FUNCTION "Wips Have Matching Index" : Bool   // FC111, SCL
{ S7_Optimized_Access := 'TRUE' }
VERSION : 0.1
   VAR_INPUT
      selected_station_wips : Array[0.."wipCount"] of "Station: Wip: Wip Module";
      evaluation_station_wips : Array[0.."wipCount"] of "Station: Wip: Wip Module";
   END_VAR
   VAR_TEMP
      code_selected : DInt;
      code_evaluation : DInt;
      p_selected : Int;
      p_evaluation : Int;
      ret : Bool;
   END_VAR
   VAR CONSTANT
      null_value : Int := -1;
   END_VAR
BEGIN
   REGION "SCAN EACH WIP IN SELECTED STATION"
       FOR #p_selected := 0 TO "wipCount" DO

           REGION "IGNORE EMPTY WIPS"
               IF #selected_station_wips[#p_selected].wip.code <> #null_value THEN

                   REGION "SCAN EACH WIP IN EVALUATION STATION"
                       FOR #p_evaluation := 0 TO "wipCount" DO

                           REGION "SAVE CODES TO LOCAL VARIABLES"
                               #code_selected := #selected_station_wips[#p_selected].wip.code;
                               #code_evaluation := #evaluation_station_wips[#p_evaluation].wip.code;
                           END_REGION

                           REGION "COMPARE CODES"
                               IF #code_selected = #code_evaluation THEN
                                   #ret := true;
                                   EXIT;
                               END_IF;
                           END_REGION

                       END_FOR;
                   END_REGION

                   REGION "EXIT OUTER LOOP IF FOUND"
                       IF #ret THEN
                           EXIT;
                       END_IF;
                   END_REGION

               END_IF;
           END_REGION

       END_FOR;
   END_REGION


   REGION "RETURN"
       #"Wips Have Matching Index" := #ret;
   END_REGION
END_FUNCTION

FUNCTION "Modify Selectable Station List: Matching WIP" : Void   // FC112, SCL
{ S7_Optimized_Access := 'TRUE' }
VERSION : 0.1
   VAR_INPUT
      saved_wips : Array[0.."hmi_station_count"] of "WIP: Station";
      selection_change : "Station Selection Change";
      selected_stations : "Selected Stations";
   END_VAR
   VAR_IN_OUT
      selectable_stns : Array[0.."stnCount"] of Int;
      selectable_stn_cnt : Int;
      visible_stations : Array[0.."slct_stn_btn_count"] of Int;
   END_VAR
   VAR_TEMP
      has_matching_wip : Bool;
      i : Int;
      p_evaluation : Int;
      selected_station : "WIP: Station";
      selected_stations_count : Int;
      selected_stations_indices : Array[0.."stnCount"] of Int;
      station_index : Int;
      t_selectable_stns : Array[0.."stnCount"] of Int;
      t_selectable_stn_count : Int;
   END_VAR
   VAR CONSTANT
      null_value : Int := -1;
   END_VAR
BEGIN
   REGION "SET UP LOCALS"
       #t_selectable_stns := #selectable_stns;
       #t_selectable_stn_count := #selectable_stn_cnt;
       #selected_stations_count := "Count Selected Stations"(#selected_stations.stns);
       "List of Array of Bool Indices"(array_of_bool := #selected_stations.stns,
                                       list_of_indices => #selected_stations_indices);
   END_REGION


   REGION "CHECK EACH SELECTED STATION VS SELECTABLE STATIONS"
       FOR #i := 0 TO #selected_stations_count DO

           REGION "EXIT LOOP ON FIRST NULL"
               IF #selected_stations_indices[#i] = #null_value THEN
                   EXIT;
               END_IF;
           END_REGION

           REGION "GET SELECTED STATION DATA"
               #station_index := #selected_stations_indices[#i];
               #selected_station := "Get WIP Station by Global Index"(index := #station_index,
                                                                         recipe_stations := #saved_wips);
           END_REGION

           REGION "REMOVE STATIONS WITH NON-MATCHING WIP"
               FOR #p_evaluation := 0 TO "hmi_station_count" DO

                   REGION "DONT RUN IF SELECTED AND EVALUATION STATIONS MATCH"
                       IF #selected_station.pStn <> #saved_wips[#p_evaluation].pStn THEN

                           REGION "RUN IF EVALUATION STATION IS SELECTABLE"
                               IF "Is In Int Array"(array_of_int := #selectable_stns, search_term := #saved_wips[#p_evaluation].pStn) THEN

                                   REGION "REMOVE EVALUATION STATION FROM SELECTABLE LIST IF NO MATCHING WIPS"
                                       #has_matching_wip := "Wips Have Matching Index"(selected_station_wips := #selected_station.wip,
                                                                                       evaluation_station_wips := #saved_wips[#p_evaluation].wip);
                                       IF NOT #has_matching_wip THEN
                                           #t_selectable_stns[#p_evaluation] := #null_value;
                                       END_IF;
                                   END_REGION

                               END_IF;
                           END_REGION

                       END_IF;
                   END_REGION

               END_FOR;
           END_REGION

           REGION "COLLAPSE"
               "Collapse Int Array"(null_value := #null_value,
                                    int_array := #t_selectable_stns);
           END_REGION

       END_FOR;
   END_REGION


   REGION "GET COUNT"
       #t_selectable_stn_count := "Count Collapsed Int Array"(null_value := #null_value,
                                                              array := #t_selectable_stns);
   END_REGION


   REGION "RETURN"
       #selectable_stns := #t_selectable_stns;
       #selectable_stn_cnt := #t_selectable_stn_count;
       "Remap Int Array"(source_int_array := #t_selectable_stns,
                         destination_int_array := #visible_stations);

   END_REGION
END_FUNCTION

FUNCTION "Pop Up: Select Stations: Animations" : Void   // FC119, SCL
{ S7_Optimized_Access := 'TRUE' }
VERSION : 0.1
   VAR_INPUT
      all_stations : "Station: All Stations";
      selectable_stn_cnt : Int;
      selected_stns : "Selected Stations";
      visable_stns : Array[0.."slct_stn_btn_count"] of Int;
   END_VAR
   VAR_IN_OUT
      interface : "Select Station";
   END_VAR
   VAR_TEMP
      i : Int;
      t_interface : "Select Station";
   END_VAR
BEGIN
   REGION "COPY TO LOCAL"
       #t_interface := #interface;
   END_REGION


   REGION "ANIMATE CLOSE SCREEN BUTTON"
       #t_interface.close_screen.animate := "Animate Bool"(colorTrue := "BgLGr",
                                                           colorFalse := "BgLRd",
                                                           evalSignal := #t_interface.close_screen.actuate);
   END_REGION


   REGION "ANIMATE STATION SELECT BUTTONS"

       REGION "ACTUATE"
           FOR #i := 0 TO "slct_stn_btn_count" DO
               IF #visable_stns[#i] <> -1 THEN

                   REGION "NOT SELECTED"
                       IF NOT #selected_stns.stns[#visable_stns[#i]] THEN
                           #t_interface.stn_select_btns[#i].animate := "Animate Bool"(colorTrue := "BgLGr",
                                                                                      colorFalse := "BgGray",
                                                                                      evalSignal := #t_interface.stn_select_btns[#i].actuate);
                       END_IF;
                   END_REGION

                   REGION "SELECTED"
                       IF #selected_stns.stns[#visable_stns[#i]] THEN
                           #t_interface.stn_select_btns[#i].animate := "Animate Bool"(colorTrue := "BgLGr",
                                                                                      colorFalse := "BgLBl",
                                                                                      evalSignal := #t_interface.stn_select_btns[#i].actuate);
                       END_IF;
                   END_REGION

               END_IF;
           END_FOR;
       END_REGION

       REGION "ENABLE"
           FOR #i := 0 TO "slct_stn_btn_count" DO
               #t_interface.stn_select_btns[#i].enable := "Select Station Button Activation"(btn_index := #i,
                                                                                             selectable_stn_cnt := #selectable_stn_cnt);
           END_FOR;
       END_REGION

       REGION "VISIBLE"
           FOR #i := 0 TO "slct_stn_btn_count" DO
               #t_interface.stn_select_btns[#i].visible := "Select Station Button Activation"(btn_index := #i,
                                                                                              selectable_stn_cnt := #selectable_stn_cnt);
           END_FOR;
       END_REGION

       REGION "DISABLED"
           FOR #i := 0 TO "slct_stn_btn_count" DO
               #t_interface.stn_select_btns[#i].enable := TRUE;
           END_FOR;
           FOR #i := #selectable_stn_cnt TO "slct_stn_btn_count" DO
               #t_interface.stn_select_btns[#i].enable := FALSE;
           END_FOR;
       END_REGION

       REGION "POPULATE STATION NAMES"
           FOR #i := 0 TO "slct_stn_btn_count" DO
               IF #visable_stns[#i] <> -1 THEN
                   #t_interface.stn_select_btns[#i].label := "Populate Station Name"(lines := 2,
                                                                                     stn := #all_stations.stn[#visable_stns[#i]]);
               END_IF;
           END_FOR;
       END_REGION

   END_REGION


   REGION "ANIMATE NAV BAR"

       REGION "NOTES"
           // mapping is necessary because hmi faceplate data structures
           // cannot consist of embedded udts
       END_REGION

       REGION "MAP HMI TO PLC"
           "Nav Bar Data Map: HMI to PLC"(hmi := #t_interface.nav_bar_HMI,
                                          plc := #t_interface.nav_Bar_PLC);
       END_REGION

       REGION "ANIMATION CALLS"
           "Select Station Nav Bar Button Animation"(selectable_stations := #selectable_stn_cnt,
                                                     visible_rows := "slct_stn_btn_count",
                                                     button := #t_interface.nav_Bar_PLC.top);
           "Select Station Nav Bar Button Animation"(selectable_stations := #selectable_stn_cnt,
                                                     visible_rows := "slct_stn_btn_count",
                                                     button := #t_interface.nav_Bar_PLC.pageUp);
           "Select Station Nav Bar Button Animation"(selectable_stations := #selectable_stn_cnt,
                                                     visible_rows := "slct_stn_btn_count",
                                                     button := #t_interface.nav_Bar_PLC.lineUp);
           "Select Station Nav Bar Button Animation"(selectable_stations := #selectable_stn_cnt,
                                                     visible_rows := "slct_stn_btn_count",
                                                     button := #t_interface.nav_Bar_PLC.lineDown);
           "Select Station Nav Bar Button Animation"(selectable_stations := #selectable_stn_cnt,
                                                     visible_rows := "slct_stn_btn_count",
                                                     button := #t_interface.nav_Bar_PLC.pageDown);
           "Select Station Nav Bar Button Animation"(selectable_stations := #selectable_stn_cnt,
                                                     visible_rows := "slct_stn_btn_count",
                                                     button := #t_interface.nav_Bar_PLC.bottom);
       END_REGION

       REGION "MAP PLC TO HMI"
           "Nav Bar Data Map: PLC to HMI"(plc := #t_interface.nav_Bar_PLC,
                                          hmi := #t_interface.nav_bar_HMI);
       END_REGION

   END_REGION


   REGION "DRAW"
       #interface := #t_interface;
   END_REGION
END_FUNCTION

// folder: HMI: Warehouse/Pop Ups/Select WIP

FUNCTION_BLOCK "Pop Up: Select WIPs"   // FB28, SCL
{ S7_Optimized_Access := 'TRUE' }
VERSION : 0.1
   VAR_INPUT
      stations : "Station: All Stations";
      wip_stations : Array[0.."hmi_station_count"] of "WIP: Station";
   END_VAR
   VAR_IN_OUT
      interface : "Select WIP";
      meta_data : "Setting Meta Data";
   END_VAR
   VAR
      selectable_wips_count : Int;
   END_VAR
   VAR_TEMP
      t_interface : "Select WIP";
   END_VAR
   VAR CONSTANT
      null_value : Int := -1;
   END_VAR
BEGIN
   IF #meta_data.selection_change.selection_change THEN
       IF "Is HMI Station"(#stations.stn[#meta_data.selection_change.station_index]) THEN
           "Pop Up: Select WIPs: Build Selectable List"(meta_data := #meta_data,
                                                        selected_stations := #meta_data.selected_stns,
                                                        wip_stations := #wip_stations,
                                                        stations := #stations,
                                                        selectable_wips_count := #selectable_wips_count);
       END_IF;
   END_IF;
END_FUNCTION_BLOCK

FUNCTION "Pop Up: Select WIPs: Get Matching WIPs" : Void   // FC125, SCL
{ S7_Optimized_Access := 'TRUE' }
VERSION : 0.1
   VAR_INPUT
      outer_wips : Array[0.."wipCount"] of "Station: Wip: Wip Module";
      inner_wips : Array[0.."wipCount"] of "Station: Wip: Wip Module";
   END_VAR
   VAR_IN_OUT
      selectable_wips : "Selectable Wips";
      selectable_wips_count : Int;
   END_VAR
   VAR_TEMP
      i : Int;
      j : Int;
      t_selectable_wips : "Selectable Wips";
      t_selectable_wips_count : Int;
   END_VAR
BEGIN
   REGION "COPY TO LOCAL"
       #t_selectable_wips := #selectable_wips;
       #t_selectable_wips_count := 0;
   END_REGION

   REGION "COMPARE EACH WIP CODE IN OUTER LIST ..." 
       FOR #i := 0 TO "wipCount" DO

           REGION "LEAVE LOOP ON FIRST NULL"
               IF #outer_wips[#i].wip.code = "null_value" THEN
                   EXIT;
               END_IF;
           END_REGION

           REGION "WITH EACH IN INNER LIST AND ..."
               FOR #j := 0 TO "wipCount" DO

                   REGION "COPY MATCHES"
                       IF #outer_wips[#i].wip.code = #inner_wips[#j].wip.code THEN
                           #t_selectable_wips.wips[#t_selectable_wips_count] := #outer_wips[#i].wip.code;
                           #t_selectable_wips_count += 1;
                       END_IF;
                   END_REGION

               END_FOR;
           END_REGION

       END_FOR;
   END_REGION


   REGION "RETURN"
       #selectable_wips := #t_selectable_wips;
       #selectable_wips_count := #t_selectable_wips_count;
   END_REGION
END_FUNCTION

FUNCTION "Pop Up: Select WIPs: Build Selectable List" : Void   // FC128, SCL
{ S7_Optimized_Access := 'TRUE' }
VERSION : 0.1
   VAR_INPUT
      selected_stations : "Selected Stations";
      stations : "Station: All Stations";
      wip_stations : Array[0.."hmi_station_count"] of "WIP: Station";
   END_VAR
   VAR_IN_OUT
      meta_data : "Setting Meta Data";
      selectable_wips_count : Int;
   END_VAR
   VAR_TEMP
      global_index : Int;
      inner_wip_index : Int;
      outer_wip_index : Int;
      p_outer : Int;
      p_inner : Int;
      selected_station_count : Int;
      station : "WIP: Station";
      t_selectable_wips_count : Int;
   END_VAR
BEGIN
   REGION "INITIALIZE SELECTABLE WIPS"
       "Fill DInt Array"(int_in := -1,
                         array_out => #meta_data.selectable_wips.wips);
       #t_selectable_wips_count := 0;
   END_REGION


   REGION "Count Selected Stations"
       #selected_station_count := "Count Selected Stations"(#selected_stations.stns);
   END_REGION


   REGION "SINGLE STATION SELECTION"
       IF #selected_station_count = 1 THEN
           #global_index := "Get First Selected Station"(#selected_stations.stns);
           #outer_wip_index := "Get WIP Station Index by Global Index"(wip_stations := #wip_stations,
                                                                       global_index := #global_index);
           "Pop Up: Select WIPs: Map WIP Codes"(wip_station := #wip_stations[#outer_wip_index],
                                                selectable_wips := #meta_data.selectable_wips,
                                                selectable_wip_count := #t_selectable_wips_count);
       END_IF;
   END_REGION


   REGION "MULTI STATION SELECTION"
       IF #selected_station_count > 1 THEN
           REGION "FOR EACH STATION..."
               FOR #p_outer := 0 TO "stnCount" DO

                   REGION "IF THE STATION HAS BEEN SELECTED..."
                       IF #selected_stations.stns[#p_outer] THEN

                           REGION "GET THE WIP STATION INDEX"
                               #outer_wip_index := "Get WIP Station Index by Global Index"(wip_stations := #wip_stations,
                                                                                           global_index := #p_outer);
                           END_REGION

                           REGION "FOR EACH STATION AFTER THIS STATION..."
                               FOR #p_inner := #p_outer + 1 TO "stnCount" DO

                                   REGION "IF THE STATION HAS BEEN SELECTED"
                                       IF #selected_stations.stns[#p_inner] THEN

                                           REGION "GET THE WIP STATION INDEX"
                                               #inner_wip_index := "Get WIP Station Index by Global Index"(wip_stations := #wip_stations,
                                                                                                           global_index := #p_inner);
                                           END_REGION

                                           REGION "INSERT INTO SELECTABLE WIP ARRAY"
                                               "Pop Up: Select WIPs: Get Matching WIPs"(outer_wips := #wip_stations[#outer_wip_index].wip,
                                                                                        inner_wips := #wip_stations[#inner_wip_index].wip,
                                                                                        selectable_wips := #meta_data.selectable_wips,
                                                                                        selectable_wips_count := #t_selectable_wips_count);
                                           END_REGION

                                       END_IF;
                                   END_REGION

                               END_FOR;
                           END_REGION

                       END_IF;
                   END_REGION

               END_FOR;
           END_REGION
       END_IF;
   END_REGION


   REGION "RETURN"
       #selectable_wips_count := #t_selectable_wips_count;
   END_REGION
END_FUNCTION

FUNCTION "Pop Up: Select WIPs: Map WIP Codes" : Void   // FC129, SCL
{ S7_Optimized_Access := 'TRUE' }
VERSION : 0.1
   VAR_INPUT
      wip_station : "WIP: Station";
   END_VAR
   VAR_IN_OUT
      selectable_wips : "Selectable Wips";
      selectable_wip_count : Int;
   END_VAR
   VAR_TEMP
      i : Int;
      t_selectable_wips : "Selectable Wips";
      t_selectable_wip_count : Int;
   END_VAR
BEGIN
   REGION "COPY TO LOCAL"
       #t_selectable_wips := #selectable_wips;
       #t_selectable_wip_count := #selectable_wip_count;
   END_REGION


   REGION "MAP VALUES"
       FOR #i := 0 TO "wipCount" DO
           IF #wip_station.wip[#i].wip.code = "null_value" THEN
               EXIT;
           END_IF;
           #t_selectable_wips.wips[#i] := #wip_station.wip[#i].wip.code;
       END_FOR;
   END_REGION


   REGION "COUNT SELECTABLE WIPS"
       #t_selectable_wip_count := "Count Collapsed DInt Array"(null_value := INT_TO_DINT("null_value"),
                                                               array := #t_selectable_wips.wips);
   END_REGION


   REGION "RETURN"
       #selectable_wips := #t_selectable_wips;
       #selectable_wip_count := #t_selectable_wip_count;
   END_REGION
END_FUNCTION

// folder: HMI: Warehouse/RSP Simulation

FUNCTION_BLOCK "Sim: from Global"   // FB26, SCL
{ S7_Optimized_Access := 'TRUE' }
VERSION : 0.1
   VAR_INPUT
      stns : "Station: All Stations";
   END_VAR
   VAR_IN_OUT
      simStations : "Simulated Stations";
   END_VAR
   VAR
      old : Struct
         nextGrp : Bool;
         prevGrp : Bool;
      END_STRUCT;
   END_VAR
   VAR_TEMP
      animate : USInt;
      btnCount : Int;
      currentBtn : Bool;
      dzLabel : WString;
      firstStn : Int;
      i : Int;
      intBox : Int;
      j : Int;
      kp8Color : DWord;
      label : WString;
      oldBtn : Bool;
      pSim : Int;
      pStn : Int;
   END_VAR
   VAR CONSTANT
      space : WString := WSTRING#' ';
      lead0 : WString := WSTRING#'0';
      volvo16 : WString := WSTRING#'VOLVO 16';
   END_VAR
BEGIN
   REGION "COPY TO LOCAL"
       #firstStn := #simStations.firstStn;
   END_REGION

   REGION "RESOLVE STATION POINTER"

       REGION "PROCESS NEXT GROUP PRESS"

           REGION "COPY TO LOCAL"
               #currentBtn := #simStations.down.actuate;
               #oldBtn := #old.nextGrp;
           END_REGION

           REGION "FALLING EDGE OF NEXT GROUP"
               IF NOT #currentBtn AND #oldBtn THEN

                   REGION "INCREMENT FIRST STATION"
                       #firstStn += "simKP8Count";
                   END_REGION

                   REGION "UPPER LIMIT ROLL OVER"
                       IF #firstStn > "stnCount" THEN
                           #firstStn -= "stnCount" + 1;
                       END_IF;
                   END_REGION

               END_IF;
           END_REGION

           REGION "NEXT GROUP CHANGE DETECTION"
               #old.nextGrp := #currentBtn;
           END_REGION

       END_REGION

       REGION "PROCESS PREVIOUS GROUP PRESS"

           REGION "COPY TO LOCAL"
               #currentBtn := #simStations.up.actuate;
               #oldBtn := #old.prevGrp;
           END_REGION

           REGION "FALLING EDGE OF PREVIOUS GROUP"
               IF NOT #currentBtn AND #oldBtn THEN

                   REGION "DECREMENT FIRST STATION"
                       #firstStn -= "simKP8Count";
                   END_REGION

                   REGION "LOWER LIMIT ROLL OVER"
                       IF #firstStn < 0 THEN
                           #firstStn += "stnCount" + 1;
                       END_IF;
                   END_REGION

               END_IF;
           END_REGION

           REGION "PREVIOUS GROUP CHANGE DETECTION"
               #old.prevGrp := #currentBtn;
           END_REGION

       END_REGION

   END_REGION

   REGION "FOR EACH BUTTON"
       FOR #i := 0 TO 11 DO

           REGION "CALCULATE POINTER"
               #pStn := #i + #firstStn;
               #pSim := #i;
           END_REGION

           REGION "UPPER LIMIT ROLL OVER"
               IF #pStn > "stnCount" THEN
                   #pStn := #firstStn + #i - "stnCount" - 1;
               END_IF;
           END_REGION

           REGION "COPY TO LOCAL"
               #kp8Color := #stns.stn[#pStn].wipCmpts.ioData.kp8.tempOut;
           END_REGION

           REGION "LABEL STATIONS"

               REGION "DETERMINE LINE LABEL"
                   #label := #stns.stn[#pStn].id.lineName;
                   IF #label = #volvo16 THEN
                       #label := WSTRING#'V16';
                   END_IF;
               END_REGION

               REGION "DETERMINE DROP ZONE LABEL"
                   #intBox := USINT_TO_INT(#stns.stn[#pStn].id.dropZone);
                   IF #intBox <= 9 THEN
                       #dzLabel := CONCAT_WSTRING(IN1 := #lead0,
                                                  IN2 := "Strip Sign"(INT_TO_WSTRING(#intBox)));
                   END_IF;
                   IF #intBox >= 10 THEN
                       #dzLabel := "Strip Sign"(INT_TO_WSTRING(#intBox));
                   END_IF;
               END_REGION

               REGION "WRITE LABEL"
                   #label := CONCAT_WSTRING(IN1 := #label,
                                            IN2 := #space,
                                            IN3 := #dzLabel);
                   #simStations.me[#pSim].stn.label := #label;
               END_REGION

           END_REGION

           REGION "ANIMATE STATION LABEL"
               #simStations.me[#pSim].stn.animate := "BgGray";
           END_REGION

           REGION "FOR EACH BUTTON"
               FOR #j := 0 TO "btnCount" DO

                   REGION "COLOR BUTTONS"
                       #animate := "KP8 Driver: HMI Emulator: Animation"(kp8Color := #kp8Color,
                                                                btnNumber := #j);
                       #simStations.me[#pSim].btn.animate[#j] := #animate;
                   END_REGION

                   REGION "WRITE BUTTON LABELS"
                       #intBox := "Pointer Calc: KP8 Labels"(#j);
                       #label := "Strip Sign"(INT_TO_WSTRING(#intBox));
                       #simStations.me[#pSim].btn.labels[#j] := #label;
                   END_REGION

               END_FOR;
           END_REGION

       END_FOR;
   END_REGION

   REGION "SAVE FIRST STATION"
       #simStations.firstStn := #firstStn;
   END_REGION

   REGION "ANIMATE NEXT GROUP PRESS"
       #simStations.down.animate := "Animate Bool"(colorTrue := "BgLGr",
                                                   colorFalse := "BgGray",
                                                   evalSignal := #simStations.down.actuate);
   END_REGION

   REGION "ANIMATE PREV GROUP PARESS"
       #simStations.up.animate := "Animate Bool"(colorTrue := "BgLGr",
                                                 colorFalse := "BgGray",
                                                 evalSignal := #simStations.up.actuate);
   END_REGION
END_FUNCTION_BLOCK

FUNCTION "Sim: to Global" : Void   // FC23, SCL
{ S7_Optimized_Access := 'TRUE' }
VERSION : 0.1
   VAR_INPUT
      simStns : "Simulated Stations";
   END_VAR
   VAR_IN_OUT
      stations : "Station: All Stations";
   END_VAR
   VAR_TEMP
      i : Int;
      j : Int;
      pSim : Int;
      pStn : Int;
   END_VAR
BEGIN
   REGION "COPY TO LOCAL"
       // #btnCount := "btnCount";
       // #firstStn := #simStns.firstStn;
       // #simKP8Count := "simKP8Count";
       // #stnCount := "stnCount";
   END_REGION

   REGION "FOR EACH STATION"
       FOR #i := 0 TO "simKP8Count" DO

           REGION "CALCULATE POINTER"
               #pStn := #i + #simStns.firstStn;
               #pSim := #i;
           END_REGION

           REGION "UPPER LIMIT ROLL OVER"
               IF #pStn > "stnCount" THEN
                   #pStn := #simStns.firstStn + #i - "stnCount" - 1;
               END_IF;
           END_REGION

           REGION "COPY SIMULATED PRESSES"
               #stations.stn[#pStn].wipCmpts.ioData.kp8.input.%B1 := #simStns.me[#pSim].btn.actuate;
           END_REGION

       END_FOR;
   END_REGION
END_FUNCTION

FUNCTION "Sim: KP8 Animations" : Word   // FC84, SCL
{ S7_Optimized_Access := 'TRUE' }
VERSION : 0.1
   VAR_INPUT
      pbs : DWord;
   END_VAR
   VAR_TEMP
      ret : Word;
   END_VAR
BEGIN
   #"Sim: KP8 Animations".%B1 := #pbs.%B0;
   #"Sim: KP8 Animations".%B0 := #pbs.%B1;
END_FUNCTION

// folder: OBs

ORGANIZATION_BLOCK "Rack or station failure"   // OB86, LAD, RackStationFailure
{ S7_Optimized_Access := 'TRUE' }
VERSION : 0.1
   VAR_INPUT
      LADDR : Hw_Device;   // Hardware identifier
      Event_Class : Byte;   // Event class
      Fault_ID : Byte;   // Fault identifier
   END_VAR
BEGIN
END_ORGANIZATION_BLOCK

ORGANIZATION_BLOCK "Startup"   // OB100, LAD, Startup
TITLE = "Complete Restart"
{ S7_Optimized_Access := 'TRUE' }
VERSION : 0.1
   VAR_INPUT
      LostRetentive : Bool;   // True if retentive data are lost
      LostRTC : Bool;   // True if date and time are lost
   END_VAR
BEGIN

REGION Network 1 (SCL): HMI STATION INITIALIZATION
   "HMI Station Initialization"();
END_REGION
END_ORGANIZATION_BLOCK

ORGANIZATION_BLOCK "Programming error"   // OB121, LAD, ProgrammingError
{ S7_Optimized_Access := 'TRUE' }
VERSION : 0.1
   VAR_INPUT
      BlockNr : UInt;   // Number of causing block
      Reaction : USInt;   // 0:ignore, 1:substitute, 2:skip
      Fault_ID : Byte;   // Fault identifier
      BlockType : USInt;   // 16#01:OB, 16#02:FC, 16#03:FB, 16#04:SFC, 16#05:SFB, 16#06:DB: Type of block causing the error
      Area : USInt;   // Area where the error occured
      DBNr : DB_ANY;   // DB number if Area = DB or DI
      Csg_OBNr : OB_Any;   // Number of OB causing the error
      Csg_Prio : USInt;   // Priority of OB causing the error
      Width : USInt;   // 0:bit, 1:byte, 2:word, 3:dword, 4:lword
   END_VAR
BEGIN
END_ORGANIZATION_BLOCK

ORGANIZATION_BLOCK "IO access error"   // OB122, LAD, IOAccessError
{ S7_Optimized_Access := 'TRUE' }
VERSION : 0.1
   VAR_INPUT
      BlockNr : UInt;   // Number of causing block
      Reaction : USInt;   // 0:ignore, 1:substitute, 2:skip
      Fault_ID : Byte;   // 16#42:reading, 16#43:writing
      BlockType : USInt;   // 16#01:OB, 16#02:FC, 16#03:FB, 16#04:SFC, 16#05:SFB, 16#06:DB: Type of block causing the error
      Area : USInt;   // 16#81:I, 16#82:Q: IO area where the IOaccess error occured
      DBNr : DB_ANY;   // Reserved for system
      Csg_OBNr : OB_Any;   // Number of OB causing the error
      Csg_Prio : USInt;   // Priority of OB causing the error
      Width : USInt;   // 0:bit, 1:byte, 2:word, 3:dword, 4:lword
   END_VAR
BEGIN
END_ORGANIZATION_BLOCK

// folder: Order/States

FUNCTION_BLOCK "Order State"   // FB2, SCL
{ S7_Optimized_Access := 'TRUE' }
VERSION : 0.1
   VAR_INPUT
      pnLib : "Recipe: PN Text Library";
   END_VAR
   VAR_IN_OUT
      stns : "Station: All Stations";
   END_VAR
   VAR_TEMP
      pStn : Int;
      pBtn : Int;
      stn : "Station: Single Station";
   END_VAR
BEGIN
   REGION "FOR EACH STATION"
       FOR #pStn := 0 TO "stnCount" DO

           REGION "FOR EACH BUTTON"
               FOR #pBtn := 0 TO "btnCount" DO

                   REGION "POPULATE CURRENT STATION"
                       #stn := #stns.stn[#pStn];
                   END_REGION

                   REGION "INITIALIZE STATE"
                       "Order State: Initialize State"(newParams := #stn.wipCmpts.flags.newPN,
                                                       pnGood := #stn.wipCmpts.flags.pnGood[#pBtn],
                                                       state := #stn.wipCmpts.orderState[#pBtn]);
                   END_REGION

                   REGION "ENTER IDLE"
                       "Order State: Enter Idle"(btnFalling := #stn.wipCmpts.kp8Logical.falling.btn[#pBtn],
                                                 state := #stn.wipCmpts.orderState[#pBtn]);
                   END_REGION

                   REGION "ENTER REQUESTED"
                       "Order State: Enter Requested"(btnRising := #stn.wipCmpts.kp8Logical.rising.btn[#pBtn],
                                                      state := #stn.wipCmpts.orderState[#pBtn]);
                   END_REGION

                   REGION "ENTER REQUESTED CRITICAL"
                       "Order State: Enter Requested Critical"(timerVal := #stn.wipCmpts.timers.remaining[#pBtn],
                                                               state := #stn.wipCmpts.orderState[#pBtn]);
                   END_REGION

                   REGION "ENTER REQUESTED EXPIRED"
                       "Order State: Enter Requested Expired"(timerVal := #stn.wipCmpts.timers.remaining[#pBtn],
                                                              state := #stn.wipCmpts.orderState[#pBtn]);
                   END_REGION

                   REGION "SAVE CURRENT STATION"
                       #stns.stn[#pStn] := #stn;
                   END_REGION

               END_FOR;
           END_REGION

       END_FOR;
   END_REGION
END_FUNCTION_BLOCK

FUNCTION "Order State: Enter Idle" : Void   // FC6, SCL
{ S7_Optimized_Access := 'TRUE' }
VERSION : 0.1
   VAR_INPUT
      btnFalling : Bool;
   END_VAR
   VAR_IN_OUT
      state : Int;
   END_VAR
BEGIN
   IF #btnFalling THEN
       #state := "idle";
   END_IF;
END_FUNCTION

FUNCTION "Order State: Enter Requested" : Void   // FC7, SCL
{ S7_Optimized_Access := 'TRUE' }
VERSION : 0.1
   VAR_INPUT
      btnRising : Bool;
   END_VAR
   VAR_IN_OUT
      state : Int;
   END_VAR
BEGIN
   IF #state = "idle" THEN
       IF #btnRising THEN
           #state := "requested";
       END_IF;
   END_IF;
END_FUNCTION

FUNCTION "Order State: Initialize State" : Void   // FC10, SCL
{ S7_Optimized_Access := 'TRUE' }
VERSION : 0.1
   VAR_INPUT
      newParams : Bool;
      pnGood : Bool;
   END_VAR
   VAR_IN_OUT
      state : Int;
   END_VAR
BEGIN
   REGION "ON NEW PARAMETERS"
       IF #newParams THEN

           REGION "ON VALID PN" 
               IF #pnGood THEN

                   REGION "INITIALIZE STATE"
                       #state := BOOL_TO_INT(#pnGood);
                   END_REGION

               END_IF;
           END_REGION

       END_IF;
   END_REGION
END_FUNCTION

FUNCTION "Order State: Enter Requested Critical" : Void   // FC16, SCL
{ S7_Optimized_Access := 'TRUE' }
VERSION : 0.1
   VAR_INPUT
      timerVal : Real;
   END_VAR
   VAR_IN_OUT
      state : Int;
   END_VAR
   VAR_TEMP
      temp : Real;
   END_VAR
BEGIN
   IF #state = "requested" THEN
       IF #timerVal > 0.0 AND #timerVal <= "tCritical" THEN
           #state := "requestedCrit";
       END_IF;
   END_IF;
END_FUNCTION

FUNCTION "Order State: Enter Requested Expired" : Void   // FC17, SCL
{ S7_Optimized_Access := 'TRUE' }
VERSION : 0.1
   VAR_INPUT
      timerVal : Real;
   END_VAR
   VAR_IN_OUT
      state : Int;
   END_VAR
BEGIN
   IF #state = "requestedCrit" THEN
       IF #timerVal <= -0.001 THEN
           #state := "requestedExp";
       END_IF;
   END_IF;
END_FUNCTION

// folder: Order/Timers

FUNCTION_BLOCK "Order Timer"   // FB6, SCL
{ S7_Optimized_Access := 'TRUE' }
VERSION : 0.1
   VAR_INPUT
      pnLib : "Recipe: PN Text Library";
   END_VAR
   VAR_IN_OUT
      stns : "Station: All Stations";
   END_VAR
   VAR
      rt : "Runtime Data";
   END_VAR
   VAR_TEMP
      pStn : Int;
      pBtn : Int;
   END_VAR
BEGIN
   REGION "RUNTIME CALL"
       #rt.elapsed := RUNTIME(#rt.mem);
       #rt.asReal := LREAL_TO_REAL(#rt.elapsed);
   END_REGION

   REGION "FOR EACH STATION"
       FOR #pStn := 0 TO "stnCount" DO

           REGION "FOR EACH BUTTON"
               FOR #pBtn := 0 TO "btnCount" DO

                   REGION "INITIALIZE TIMERS"
                       "Order Timer: Initialize"(pnLib := #pnLib,
                                                 pBtn := #pBtn,
                                                 stn := #stns.stn[#pStn]);
                   END_REGION

                   REGION "EXECUTE TIMERS"
                       "Order Timer: Timer Execution"(elapsedTime := #rt.asReal,
                                                      pBtn := #pBtn,
                                                      stn:=#stns.stn[#pStn],
                                                      timers := #stns.stn[#pStn].wipCmpts.timers);
                   END_REGION

               END_FOR;
           END_REGION

       END_FOR;
   END_REGION
END_FUNCTION_BLOCK

FUNCTION "Order Timer: Initialize" : Void   // FC8, SCL
{ S7_Optimized_Access := 'TRUE' }
VERSION : 0.1
   VAR_INPUT
      pnLib : "Recipe: PN Text Library";
      pBtn : Int;
   END_VAR
   VAR_IN_OUT
      stn : "Station: Single Station";
   END_VAR
   VAR_TEMP
      pnGood : Bool;
      default : Bool;
      clear : Bool;
   END_VAR
BEGIN
   REGION "ON PN CHANGE"
       IF #stn.wipCmpts.flags.newPN THEN

           REGION "INITIALIZE TO DEFAULT"

               REGION "EXECUTION VALIDATION"
                   #default := "Order Timer: Set to Default Check"(pnGood := #stn.wipCmpts.flags.pnGood[#pBtn],
                                                                   inSettingsScreen := #stn.wipCmpts.flags.inSettingsScreen,
                                                                   timerReset := #stn.wipCmpts.flags.resetTimer[#pBtn]);
               END_REGION

               REGION "ON VALIDATION"
                   IF #default THEN

                       REGION "SET DEFAULT TIME VALUE"
                           #stn.wipCmpts.timers.ptAllotted[#pBtn] := "tAllotted";
                           #stn.wipCmpts.timers.ptCritical[#pBtn] := "tCritical";
                       END_REGION

                   END_IF;
               END_REGION

           END_REGION

           REGION "INITIALIZE TO ZERO"

               REGION "EXECUTION VALIDATION"
                   #clear := "Order Timer: Set to Zero Check"(pnGood := #stn.wipCmpts.flags.pnGood[#pBtn],
                                                              inSettingsScreen := #stn.wipCmpts.flags.inSettingsScreen,
                                                              timerReset := #stn.wipCmpts.flags.resetTimer[#pBtn]);
               END_REGION

               REGION "ON VALIDATION"
                   IF #clear THEN

                       REGION "SET DEFAULT TIME VALUE"
                           #stn.wipCmpts.timers.ptAllotted[#pBtn] := 0.0;
                           #stn.wipCmpts.timers.ptCritical[#pBtn] := 0.0;
                       END_REGION

                   END_IF;
               END_REGION

           END_REGION

       END_IF;
   END_REGION
END_FUNCTION

FUNCTION "Order Timer: Timer Execution" : Void   // FC11, SCL
{ S7_Optimized_Access := 'TRUE' }
VERSION : 0.1
   VAR_INPUT
      elapsedTime : Real;
      pBtn : Int;
      stn : "Station: Single Station";
   END_VAR
   VAR_IN_OUT
      timers : "Station: Timers";
   END_VAR
BEGIN
   REGION "RUN CONDITIONS"
       CASE #stn.wipCmpts.orderState[#pBtn] OF

           "reset", "idle":
               IF #stn.flags.stateTransition[#pBtn] THEN
                   #timers.elapsed[#pBtn] := 0.0;
                   #timers.remaining[#pBtn] := 0.0;
               END_IF;

           "requested".."acknowledgedExp":
               #timers.elapsed[#pBtn] += #elapsedTime;
               #timers.remaining[#pBtn] := #timers.ptAllotted[#pBtn] - #timers.elapsed[#pBtn];

           ELSE:
               ;

       END_CASE;
   END_REGION
END_FUNCTION

FUNCTION "Order Timer: Set to Default Check" : Bool   // FC12, SCL
{ S7_Optimized_Access := 'TRUE' }
VERSION : 0.1
   VAR_INPUT
      pnGood : Bool;
      inSettingsScreen : Bool;
      timerReset : Bool;
   END_VAR
   VAR_TEMP
      ret : Bool;
   END_VAR
BEGIN
   REGION "ON VALID PN"
       #ret := #pnGood;
   END_REGION

   REGION "NOT WHILE IN SETTINGS SCREEN"
       IF #inSettingsScreen THEN
           #ret := FALSE;
       END_IF;
   END_REGION

   REGION "ON RESET REQUEST"
       #ret := #timerReset OR #ret;
   END_REGION

   REGION "RETURN"
       #"Order Timer: Set to Default Check" := #ret;
   END_REGION
END_FUNCTION

FUNCTION "Order Timer: Set to Zero Check" : Bool   // FC15, SCL
{ S7_Optimized_Access := 'TRUE' }
VERSION : 0.1
   VAR_INPUT
      pnGood : Bool;
      inSettingsScreen : Bool;
      timerReset : Bool;
   END_VAR
   VAR_TEMP
      ret : Bool;
   END_VAR
BEGIN
   REGION "ON VALID PN"
       #ret := NOT #pnGood;
   END_REGION

   REGION "NOT WHILE IN SETTINGS SCREEN"
       IF #inSettingsScreen THEN
           #ret := FALSE;
       END_IF;
   END_REGION

   REGION "ON RESET REQUEST"
       #ret := #timerReset OR #ret;
   END_REGION

   REGION "RETURN"
       #"Order Timer: Set to Zero Check" := #ret;
   END_REGION
END_FUNCTION

// folder: Part Request

FUNCTION_BLOCK "Part Request"   // FB7, SCL
{ S7_Optimized_Access := 'TRUE' }
VERSION : 0.1
   VAR_INPUT
      stns : "Station: All Stations";
      savedWips : "Recipe: HMI Stations Saved Wips";
      pnLib : "Recipe: PN Text Library";
   END_VAR
   VAR_IN_OUT
      dataTable : "Part Request Data";
   END_VAR
   VAR RETAIN
      pDataRow : Int;
   END_VAR
   VAR_TEMP
      address : DInt;
      addRequest : Bool;
      inTable : DInt;
      pStn : Int;
      pBtn : Int;
      pWip : Int;
      pRqstsRow : Int;
      removeRequest : Bool;
   END_VAR
BEGIN
   REGION "FOR EACH STATION"
       FOR #pStn := 0 TO "stnCount" DO

           REGION "FOR EACH BUTTON"
               FOR #pBtn := 0 TO "btnCount" DO

                   REGION "NEXT BUTTON ON NO TRANSITION"
                       IF NOT #stns.stn[#pStn].flags.stateTransition[#pBtn] THEN
                           GOTO NOSTNREQ;
                       END_IF;
                   END_REGION

                   REGION "GET ADDRESS"
                       #pWip := DINT_TO_INT(#stns.stn[#pStn].wipData.index);
                       #address := "Address: Set Address"(pStn := #pStn, pBtn := #pBtn, pWip := #pWip);
                   END_REGION

                   REGION "CHECK FOR ENTRY IN DATA TABLE"
                       #inTable := "Part Request: Address in Table"(search := #address,
                                                                    dataTable := #dataTable);
                   END_REGION

                   REGION "ADD"

                       REGION "VALIDATE CONDITIONS"
                           #addRequest := "Part Request: Validate Add"(inTable := #inTable,
                                                                       orderState := #stns.stn[#pStn].wipCmpts.orderState[#pBtn]);
                       END_REGION

                       REGION "EXECUTE"
                           IF #addRequest THEN
                               #addRequest := FALSE;
                               #dataTable.row[#pDataRow] := #address;
                               "Row Pointer: Roll Over"(limit := "partReqDataRowCount",
                                                                "pointer" := #pDataRow);
                           END_IF;
                       END_REGION

                   END_REGION

                   REGION "REMOVE SINGLE STATION"

                       REGION "VALIDATE CONDITIONS: SINGLE"
                           #removeRequest := "Part Request: Validate Remove: Single"(inTable := #inTable,
                                                                                     orderState := #stns.stn[#pStn].wipCmpts.orderState[#pBtn]);
                       END_REGION

                       REGION "EXECUTE"
                           IF #removeRequest THEN
                               #removeRequest := FALSE;
                               #dataTable.row[#inTable] := -1;
                               "Part Request: Collapse Table"(#dataTable);
                               "Row Pointer: Post Collapse"(dataTable := #dataTable,
                                                            pDataRow := #pDataRow);
                           END_IF;
                       END_REGION

                   END_REGION

               NOSTNREQ:
                   ;
               END_FOR;
           END_REGION

       END_FOR;
   END_REGION


   (* REGION "REMOVE WIP STATIONS"                    
       FOR #pStn := 0 TO "hmiStnCount" DO
           FOR #pWip := 0 TO "wipCount" DO
               IF #savedWips.stn[#pStn].wip[#pWip].flags.clearWipRequest THEN
                   FOR #pBtn := 0 TO "btnCount" DO
                       #address := "Address: Set Address"(pBtn := #pBtn, pStn := #pStn, pWip := #pWip);
                       #inTable := "Part Request: Address in Table"(adrRequest := #address,
                                                                    dataTable := #dataTable);
                       #removeRequest := "Part Request: Validate Remove: WIP"(inTable := #inTable,
                                                                              clearWipRequest := #savedWips.stn[#pStn].wip[#pWip].flags.clearWipRequest);
                       IF #removeRequest THEN
                           #removeRequest := FALSE;
                           "Part Request: Remove"(pRow := #inTable,
                                                  dataTable := #dataTable);
                           "Part Request: Collapse Table"(#dataTable);
                           "Row Pointer: Post Collapse"(dataTable := #dataTable,
                                                        pDataRow := #pDataRow);
                       END_IF;
                   END_FOR;
               END_IF;
           END_FOR;
       END_FOR;
   END_REGION *)
END_FUNCTION_BLOCK

FUNCTION "Part Request: Address in Table" : DInt   // FC27, SCL
{ S7_Optimized_Access := 'TRUE' }
VERSION : 0.1
   VAR_INPUT
      search : DInt;
      dataTable : "Part Request Data";
   END_VAR
   VAR_TEMP
      ret : DInt;
      pRow : DInt;
   END_VAR
BEGIN
   REGION "DEFAULT RETURN"    
       #ret := -1;
   END_REGION

   REGION "CHECK TABLE"
       WHILE #dataTable.row[#pRow] <> #search AND #pRow <= "partReqDataRowCount" DO
           #pRow += 1;
       END_WHILE;
       IF #pRow <= "partReqDataRowCount" THEN
           #ret := #pRow;
       END_IF;
   END_REGION

   REGION "RETURN"
       #"Part Request: Address in Table" := #ret;
   END_REGION

   REGION "CALL READ VFD"
       ;
       ;
   END_REGION
END_FUNCTION

FUNCTION "Part Request: Validate Add" : Bool   // FC30, SCL
{ S7_Optimized_Access := 'TRUE' }
VERSION : 0.1
   VAR_INPUT
      inTable : DInt;
      orderState : Int;
   END_VAR
   VAR_TEMP
      ret : Bool;
   END_VAR
BEGIN
   IF #inTable = -1 THEN
       CASE #orderState OF
           "idle",
           "requestedCrit", "requestedExp",
           "ordered", "orderedCrit", "orderedExp",
           "acknowledged", "acknowledgedCrit", "acknowledgedExp":
               #ret := FALSE;
           "requested":
               #ret := TRUE;
       END_CASE;
   END_IF;
   #"Part Request: Validate Add" := #ret;
END_FUNCTION

FUNCTION "Part Request: Validate Remove: Single" : Bool   // FC41, SCL
{ S7_Optimized_Access := 'TRUE' }
VERSION : 0.1
   VAR_INPUT
      inTable : DInt;
      orderState : Int;
   END_VAR
   VAR_TEMP
      ret : Bool;
   END_VAR
BEGIN
   IF #inTable <> -1 THEN
       CASE #orderState OF
           "requested", "requestedCrit", "requestedExp",
           "ordered", "orderedCrit", "orderedExp",
           "acknowledged", "acknowledgedCrit", "acknowledgedExp":
               #ret := FALSE;
           "idle":
               #ret := TRUE;
       END_CASE;
   END_IF;
   #"Part Request: Validate Remove: Single" := #ret;
END_FUNCTION

FUNCTION "Part Request: Clear Data Table" : Void   // FC48, SCL
{ S7_Optimized_Access := 'TRUE' }
VERSION : 0.1
   VAR_IN_OUT
      dataTable : "Part Request Data";
   END_VAR
   VAR_TEMP
      pRow : Int;
   END_VAR
   VAR CONSTANT
      clearRow : DInt := -1;
   END_VAR
BEGIN
   FOR #pRow := 0 TO "partReqDataRowCount" DO
       #dataTable.row[#pRow] := #clearRow;
   END_FOR;
END_FUNCTION

FUNCTION "Part Request: Collapse Table" : Void   // FC55, SCL
{ S7_Optimized_Access := 'TRUE' }
VERSION : 0.1
   VAR_IN_OUT
      dataTable : "Part Request Data";
   END_VAR
   VAR_TEMP
      pRow : Int;
      pScan : Int;
   END_VAR
BEGIN
   FOR #pRow := 0 TO "partReqDataRowCount" DO
       #pScan := 1;
       IF #dataTable.row[#pRow] <= -1 THEN
           WHILE #dataTable.row[#pRow + #pScan] <= -1 AND #pRow + #pScan < "partReqDataRowCount" DO
               #pScan += 1;
           END_WHILE;
           #dataTable.row[#pRow] := #dataTable.row[#pRow + #pScan];
           #dataTable.row[#pRow + #pScan] := -1;
           IF #pRow + #pScan = "partReqDataRowCount" THEN
               RETURN;
           END_IF;
       END_IF;
   END_FOR;
END_FUNCTION

FUNCTION "Part Request: Validate Remove: WIP" : Bool   // FC89, SCL
{ S7_Optimized_Access := 'TRUE' }
VERSION : 0.1
   VAR_INPUT
      inTable : DInt;
      clearWipRequest : Bool;
   END_VAR
   VAR_TEMP
      ret : Bool;
   END_VAR
BEGIN
   IF #inTable <> -1 THEN
       #ret := #clearWipRequest;
   END_IF;

   #"Part Request: Validate Remove: WIP" := #ret;
END_FUNCTION

// folder: Stations

FUNCTION_BLOCK "Button Parameters"   // FB12, SCL
{ S7_Optimized_Access := 'TRUE' }
VERSION : 0.1
   VAR_INPUT
      pnLib : "Recipe: PN Text Library";
   END_VAR
   VAR_IN_OUT
      stns : "Station: All Stations";
   END_VAR
   VAR
      placeHolder : Bool;
   END_VAR
   VAR_TEMP
      pBtn : Int;
      pStn : Int;
   END_VAR
BEGIN
   REGION "FOR EACH STATION"
       FOR #pStn := 0 TO "stnCount" DO

           REGION "ON CODE CHANGE"
               IF #stns.stn[#pStn].wipCmpts.flags.newPN THEN

                   REGION "FOR EACH BUTTON"
                       FOR #pBtn := 0 TO "btnCount" DO

                           REGION "LOAD PARAMETERS"
                               "Load Button Parameters OP"(pnGood := #stns.stn[#pStn].wipCmpts.flags.pnGood[#pBtn],
                                                           btnConfig := #stns.stn[#pStn].kp8Config.btn[#pBtn]);
                           END_REGION

                       END_FOR;
                   END_REGION

               END_IF;
           END_REGION

       END_FOR;
   END_REGION
END_FUNCTION_BLOCK

FUNCTION "Load Button Parameters OP" : Void   // FC2, SCL
{ S7_Optimized_Access := 'TRUE' }
VERSION : 0.1
   VAR_INPUT
      pnGood : Bool;
   END_VAR
   VAR_IN_OUT
      btnConfig : "KP8 Driver: Parameters: 1 Button";
   END_VAR
BEGIN
   REGION "ON GOOD PN"
       IF #pnGood THEN

           REGION "ACTIVATE BUTTON"
               #btnConfig.activate := TRUE;
               #btnConfig.cOff := 'green';
               #btnConfig.cOn1 := 'yellow';
               #btnConfig.cOn2 := '';
               #btnConfig.flash := FALSE;
               #btnConfig.group := 0;
               #btnConfig.mode := TRUE;
           END_REGION

       END_IF;
   END_REGION